(* Logix 5000 project; controller PLC_MCC1201_220AP1 vendor 1 type 14 code 164 rev 35.11; software revision 35.00; part 14 of 25 *)
(* tags used below, declared in another part *)
   AFI : ALIAS FOR B3[7].15;
   B175 : DINT[1];
   B176 : DINT[1];
   B180 : DINT[10];
   B3 : DINT[102];
   B52 : DINT[100];
   C183 : COUNTER[3];
   C1_ACTIVE_LAMP : ALIAS FOR N54[260].0;
   C2_ACTIVE_LAMP : ALIAS FOR N54[261].0;
   C3_ACTIVE_LAMP : ALIAS FOR N54[262].0;
   C5 : COUNTER[100];
   C5_ACTIVE_LAMP : ALIAS FOR N54[264].0;
   CR1_DOWN_PROX : ALIAS FOR I[64].11;
   I : INT[128];
   LEHR_2IN_PULSE : ALIAS FOR B73[0].1;
   LEHR_SPEED : ALIAS FOR N60[1];
   LEHRSPD_CURRENT : ALIAS FOR N98[5];
   MS_ACCUM : ALIAS FOR N70[1];
   MS_LEHR : ALIAS FOR N60[11];
   MSEC_TRIM : ALIAS FOR N60[12];
   N125 : DINT[414];
   N126 : DINT[103];
   N127 : DINT[997];
   N128 : DINT[997];
   N177 : DINT[5];
   N177_0 : ALIAS FOR N177[0];
   N188 : DINT[500];
   N26 : DINT[1000];
   N54 : DINT[501];
   N70 : DINT[3];
   N80 : DINT[16];
   O : INT[128];
   RELDR_ESTOP : ALIAS FOR I[80].0;
   S : INT[128];
   T182 : TIMER[11];
   T4 : TIMER[100];
   TMP_xAlwaysOFF : BOOL;
   TONY : ALIAS FOR B3[10].15;
   TRIM_2IN_PULSE : ALIAS FOR B73[0].2;
   TRIM_SPEED : ALIAS FOR N60[2];
(* MainProgram, continued *)

ROUTINE _16_PULSER   (* ladder *)
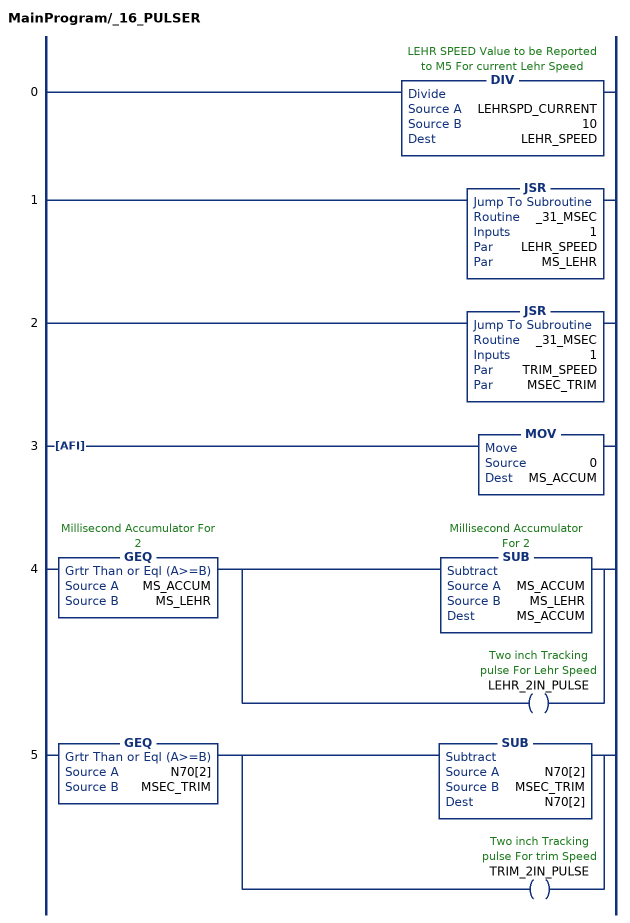
   0: DIV(LEHRSPD_CURRENT,10,LEHR_SPEED);
   1: JSR(_31_MSEC,1,LEHR_SPEED,MS_LEHR);
   2: JSR(_31_MSEC,1,TRIM_SPEED,MSEC_TRIM);
   3: AFI()MOV(0,MS_ACCUM);
   4: GEQ(MS_ACCUM,MS_LEHR)[SUB(MS_ACCUM,MS_LEHR,MS_ACCUM) ,OTE(LEHR_2IN_PULSE) ];
   5: GEQ(N70[2],MSEC_TRIM)[SUB(N70[2],MSEC_TRIM,N70[2]) ,OTE(TRIM_2IN_PULSE) ];
END_ROUTINE

ROUTINE _17_LADDER   (* ladder *)
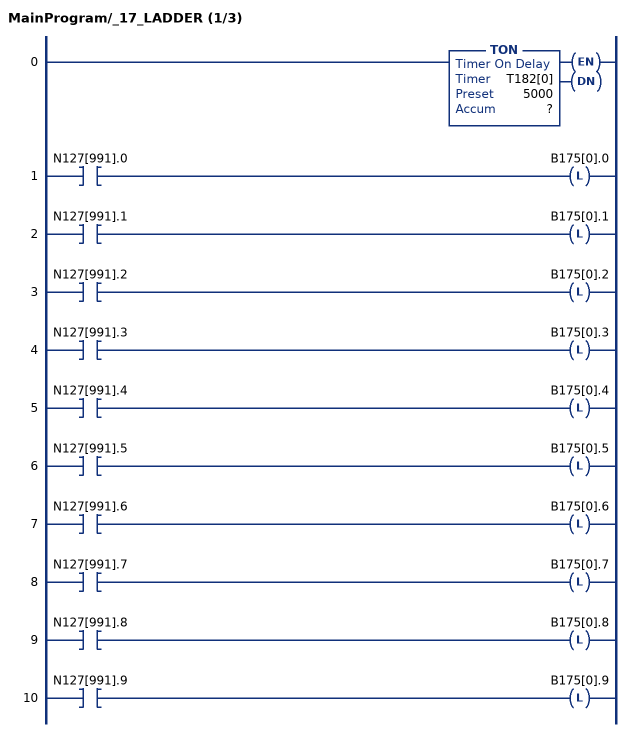
   0: TON(T182[0],?,?);
   1: XIC(N127[991].0)OTL(B175[0].0);
   2: XIC(N127[991].1)OTL(B175[0].1);
   3: XIC(N127[991].2)OTL(B175[0].2);
   4: XIC(N127[991].3)OTL(B175[0].3);
   5: XIC(N127[991].4)OTL(B175[0].4);
   6: XIC(N127[991].5)OTL(B175[0].5);
   7: XIC(N127[991].6)OTL(B175[0].6);
   8: XIC(N127[991].7)OTL(B175[0].7);
   9: XIC(N127[991].8)OTL(B175[0].8);
   10: XIC(N127[991].9)OTL(B175[0].9);
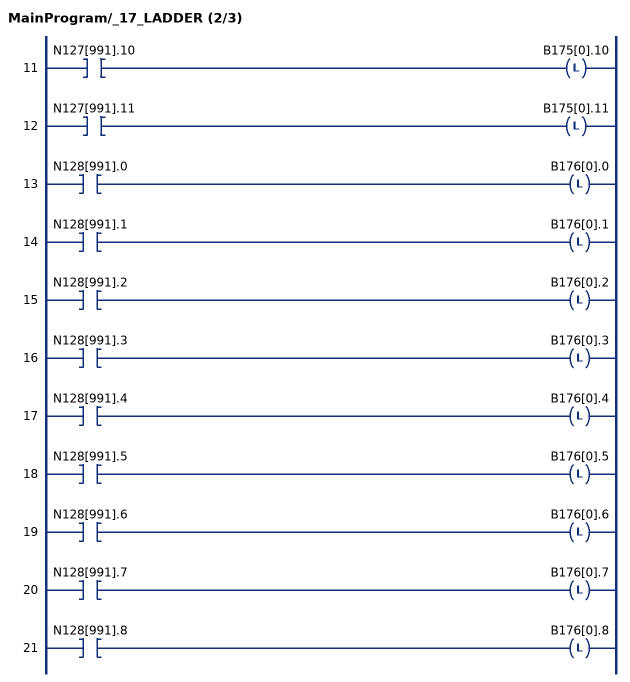
   11: XIC(N127[991].10)OTL(B175[0].10);
   12: XIC(N127[991].11)OTL(B175[0].11);
   13: XIC(N128[991].0)OTL(B176[0].0);
   14: XIC(N128[991].1)OTL(B176[0].1);
   15: XIC(N128[991].2)OTL(B176[0].2);
   16: XIC(N128[991].3)OTL(B176[0].3);
   17: XIC(N128[991].4)OTL(B176[0].4);
   18: XIC(N128[991].5)OTL(B176[0].5);
   19: XIC(N128[991].6)OTL(B176[0].6);
   20: XIC(N128[991].7)OTL(B176[0].7);
   21: XIC(N128[991].8)OTL(B176[0].8);
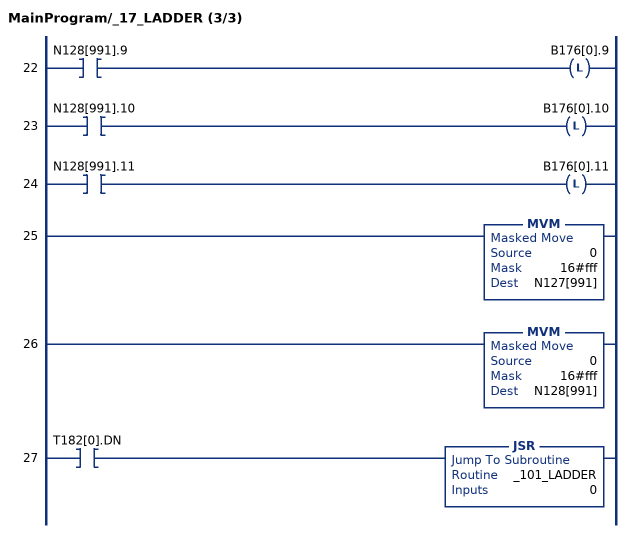
   22: XIC(N128[991].9)OTL(B176[0].9);
   23: XIC(N128[991].10)OTL(B176[0].10);
   24: XIC(N128[991].11)OTL(B176[0].11);
   25: MVM(0,16#fff,N127[991]);
   26: MVM(0,16#fff,N128[991]);
   27: XIC(T182[0].DN)JSR(_101_LADDER,0);
END_ROUTINE

ROUTINE _19_PII   (* ladder *)
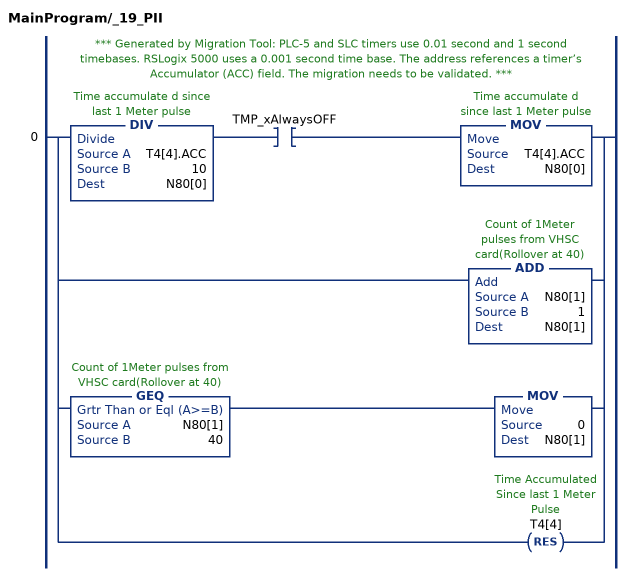
   // *** Generated by Migration Tool: PLC-5 and SLC timers use 0.01 second and 1 second timebases. RSLogix 5000 uses a 0.001 second time base. The address references a timer’s Accumulator (ACC) field. The migration needs to be validated. ***
   0: [DIV(T4[4].ACC,10,N80[0]) XIC(TMP_xAlwaysOFF) MOV(T4[4].ACC,N80[0]) ,ADD(N80[1],1,N80[1]) ,GEQ(N80[1],40) MOV(0,N80[1]) ,RES(T4[4]) ];
END_ROUTINE

ROUTINE _22_LADDER   (* ladder *)
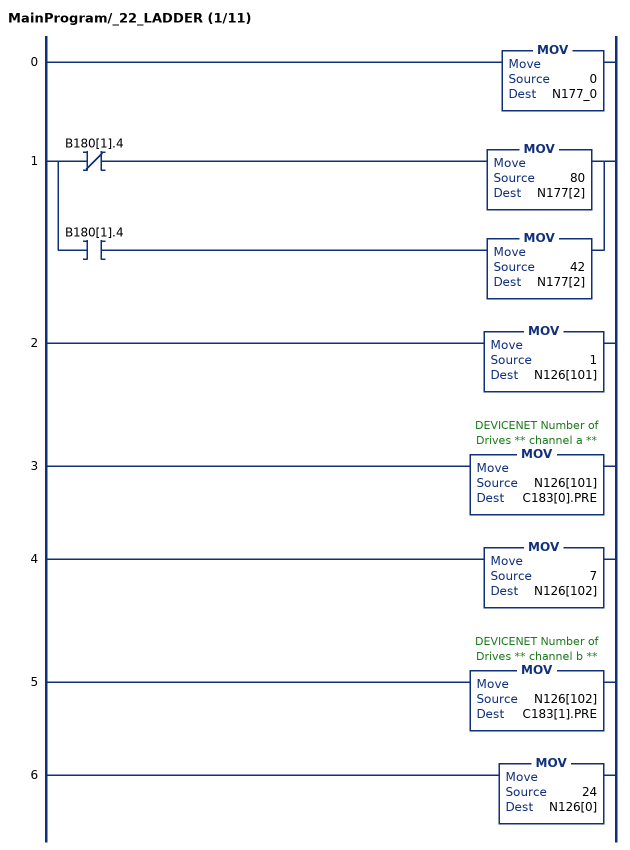
   0: MOV(0,N177_0);
   1: [XIO(B180[1].4) MOV(80,N177[2]) ,XIC(B180[1].4) MOV(42,N177[2]) ];
   2: MOV(1,N126[101]);
   3: MOV(N126[101],C183[0].PRE);
   4: MOV(7,N126[102]);
   5: MOV(N126[102],C183[1].PRE);
   6: MOV(24,N126[0]);
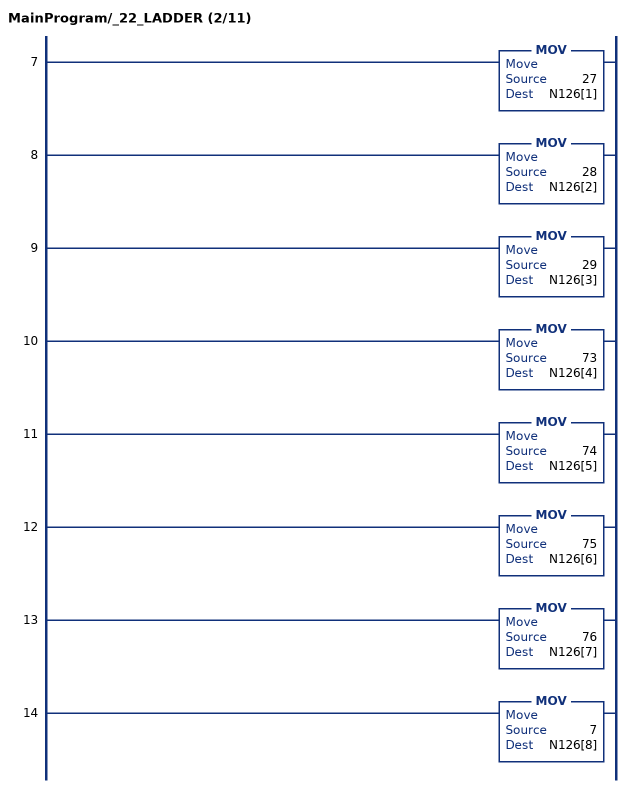
   7: MOV(27,N126[1]);
   8: MOV(28,N126[2]);
   9: MOV(29,N126[3]);
   10: MOV(73,N126[4]);
   11: MOV(74,N126[5]);
   12: MOV(75,N126[6]);
   13: MOV(76,N126[7]);
   14: MOV(7,N126[8]);
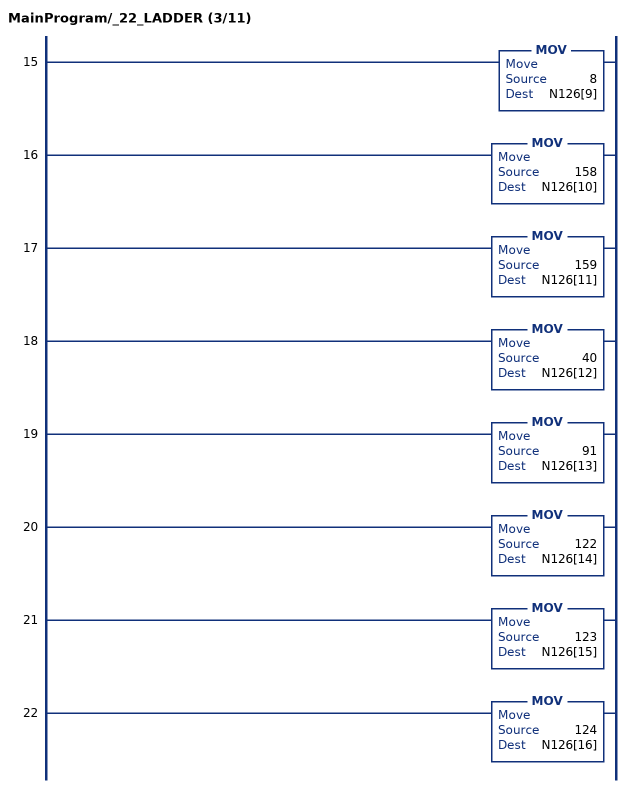
   15: MOV(8,N126[9]);
   16: MOV(158,N126[10]);
   17: MOV(159,N126[11]);
   18: MOV(40,N126[12]);
   19: MOV(91,N126[13]);
   20: MOV(122,N126[14]);
   21: MOV(123,N126[15]);
   22: MOV(124,N126[16]);
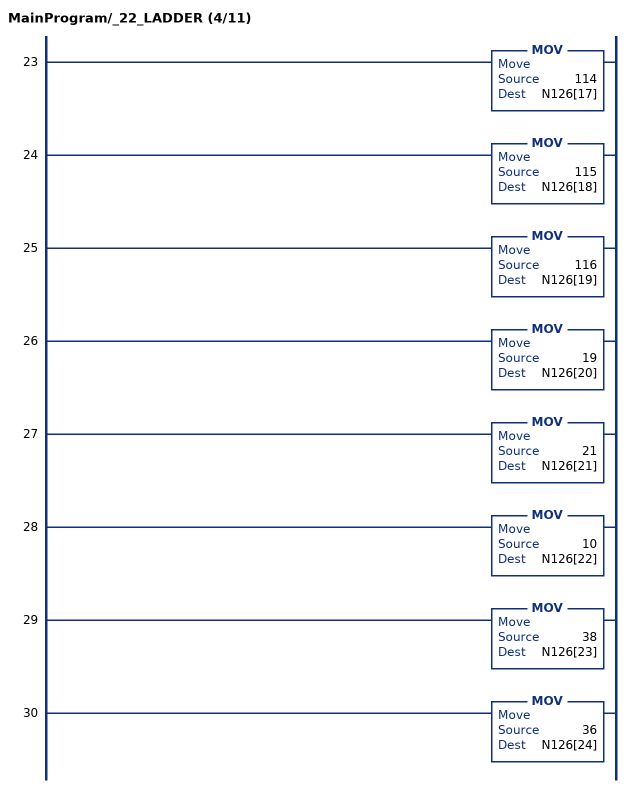
   23: MOV(114,N126[17]);
   24: MOV(115,N126[18]);
   25: MOV(116,N126[19]);
   26: MOV(19,N126[20]);
   27: MOV(21,N126[21]);
   28: MOV(10,N126[22]);
   29: MOV(38,N126[23]);
   30: MOV(36,N126[24]);
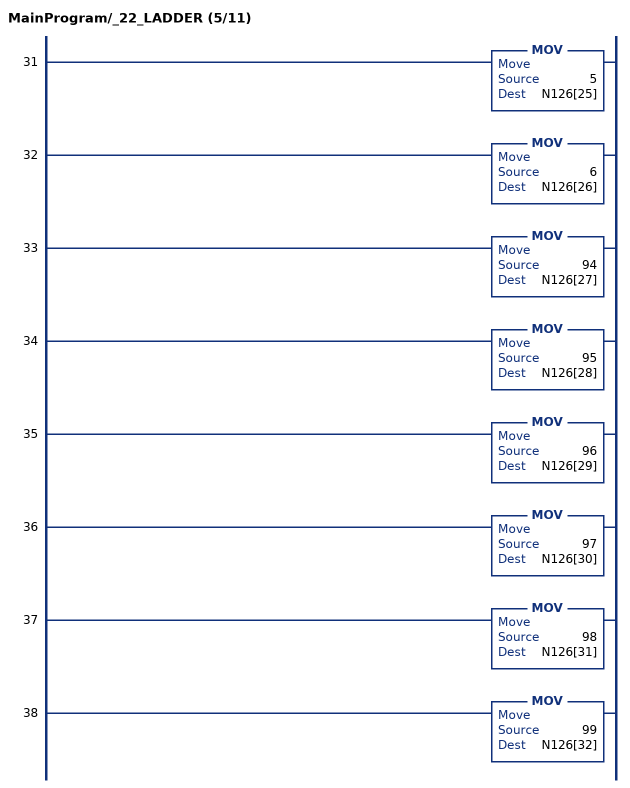
   31: MOV(5,N126[25]);
   32: MOV(6,N126[26]);
   33: MOV(94,N126[27]);
   34: MOV(95,N126[28]);
   35: MOV(96,N126[29]);
   36: MOV(97,N126[30]);
   37: MOV(98,N126[31]);
   38: MOV(99,N126[32]);
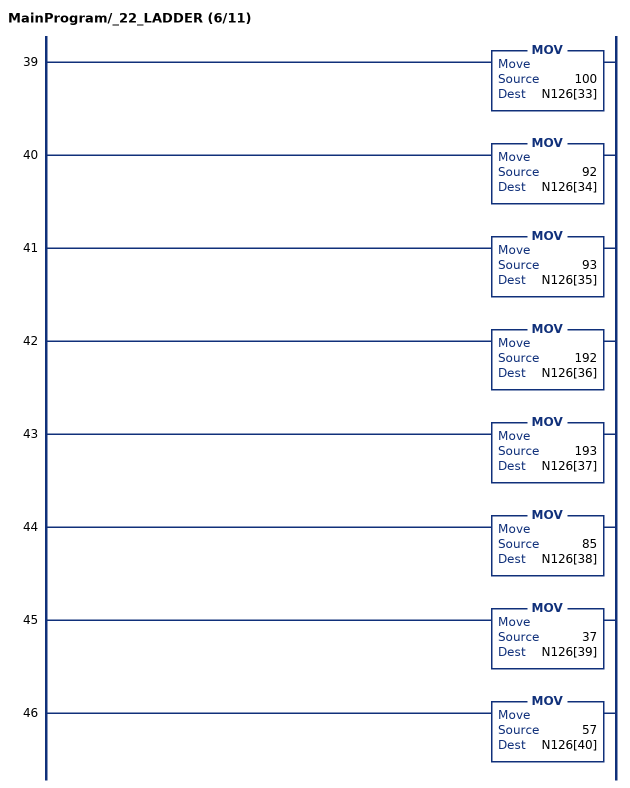
   39: MOV(100,N126[33]);
   40: MOV(92,N126[34]);
   41: MOV(93,N126[35]);
   42: MOV(192,N126[36]);
   43: MOV(193,N126[37]);
   44: MOV(85,N126[38]);
   45: MOV(37,N126[39]);
   46: MOV(57,N126[40]);
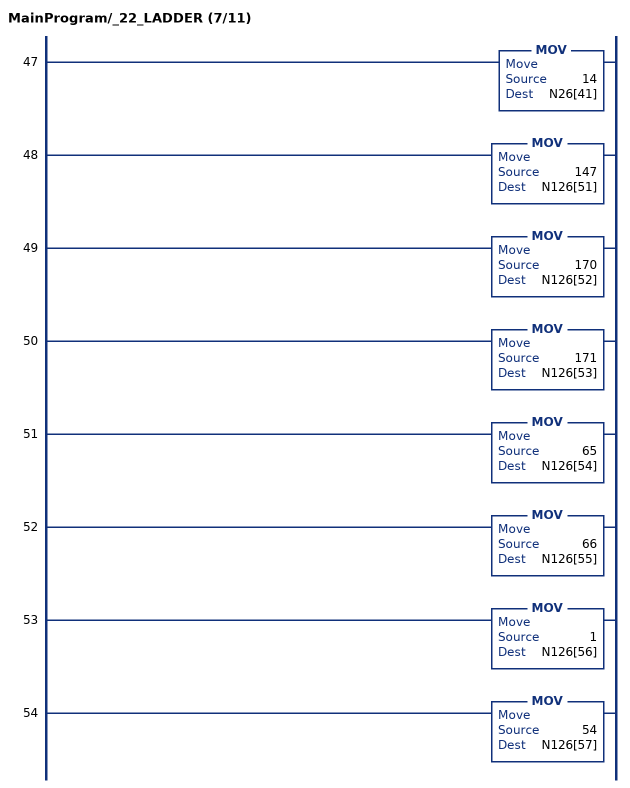
   47: MOV(14,N26[41]);
   48: MOV(147,N126[51]);
   49: MOV(170,N126[52]);
   50: MOV(171,N126[53]);
   51: MOV(65,N126[54]);
   52: MOV(66,N126[55]);
   53: MOV(1,N126[56]);
   54: MOV(54,N126[57]);
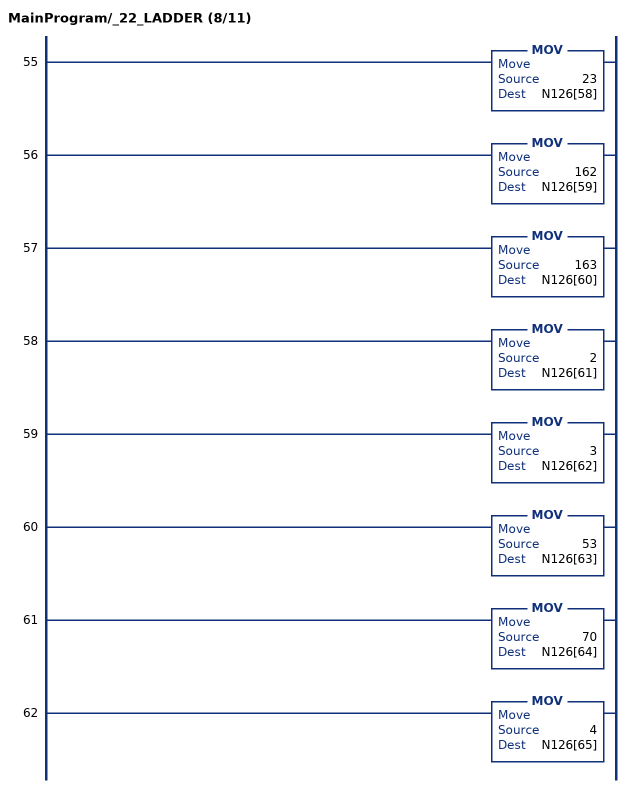
   55: MOV(23,N126[58]);
   56: MOV(162,N126[59]);
   57: MOV(163,N126[60]);
   58: MOV(2,N126[61]);
   59: MOV(3,N126[62]);
   60: MOV(53,N126[63]);
   61: MOV(70,N126[64]);
   62: MOV(4,N126[65]);
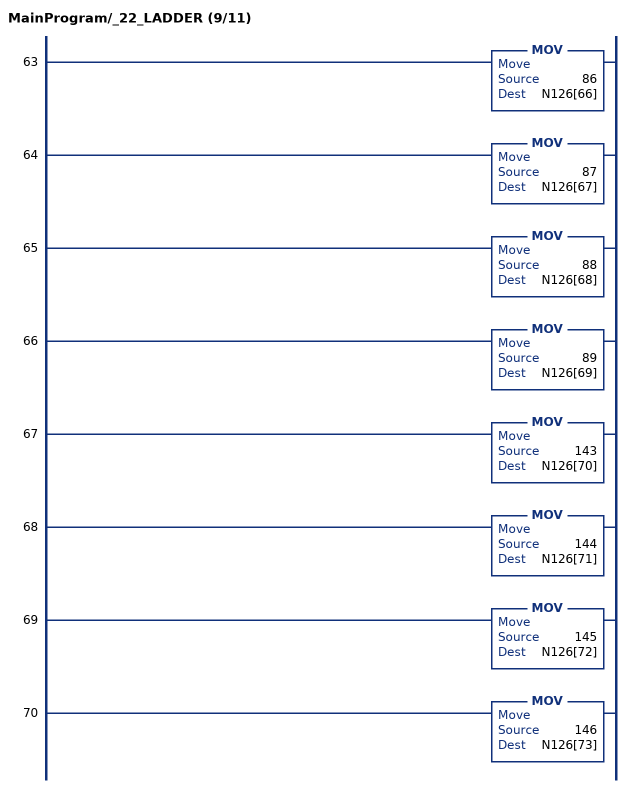
   63: MOV(86,N126[66]);
   64: MOV(87,N126[67]);
   65: MOV(88,N126[68]);
   66: MOV(89,N126[69]);
   67: MOV(143,N126[70]);
   68: MOV(144,N126[71]);
   69: MOV(145,N126[72]);
   70: MOV(146,N126[73]);
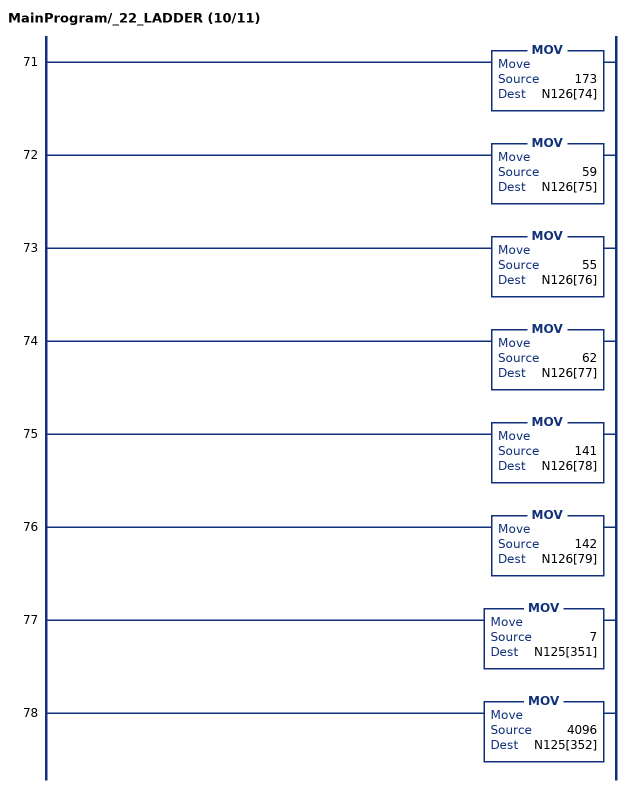
   71: MOV(173,N126[74]);
   72: MOV(59,N126[75]);
   73: MOV(55,N126[76]);
   74: MOV(62,N126[77]);
   75: MOV(141,N126[78]);
   76: MOV(142,N126[79]);
   77: MOV(7,N125[351]);
   78: MOV(4096,N125[352]);
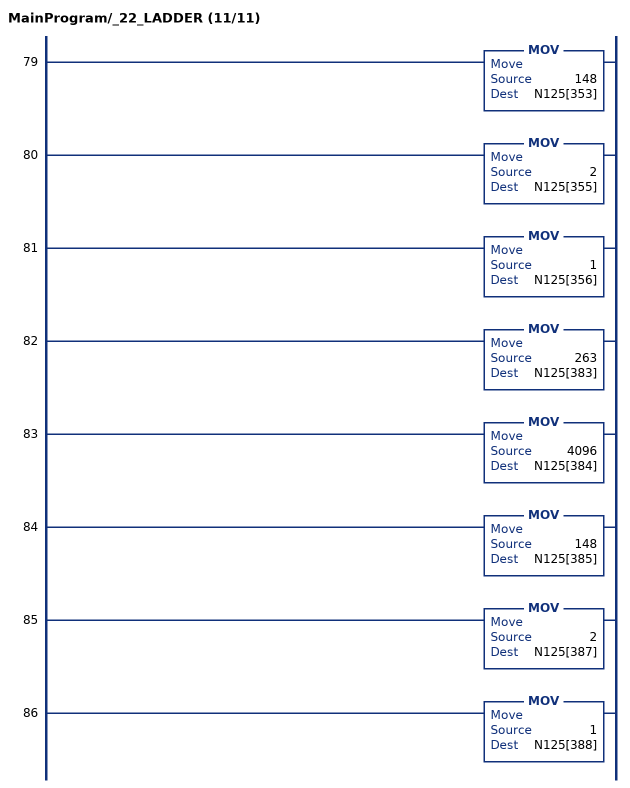
   79: MOV(148,N125[353]);
   80: MOV(2,N125[355]);
   81: MOV(1,N125[356]);
   82: MOV(263,N125[383]);
   83: MOV(4096,N125[384]);
   84: MOV(148,N125[385]);
   85: MOV(2,N125[387]);
   86: MOV(1,N125[388]);
END_ROUTINE

ROUTINE _24_ADAPTER   (* ladder *)
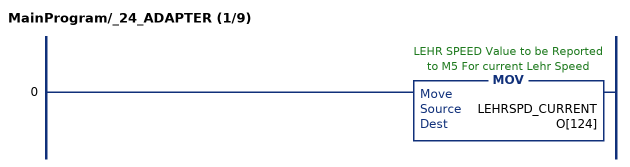
   0: MOV(LEHRSPD_CURRENT,O[124]);
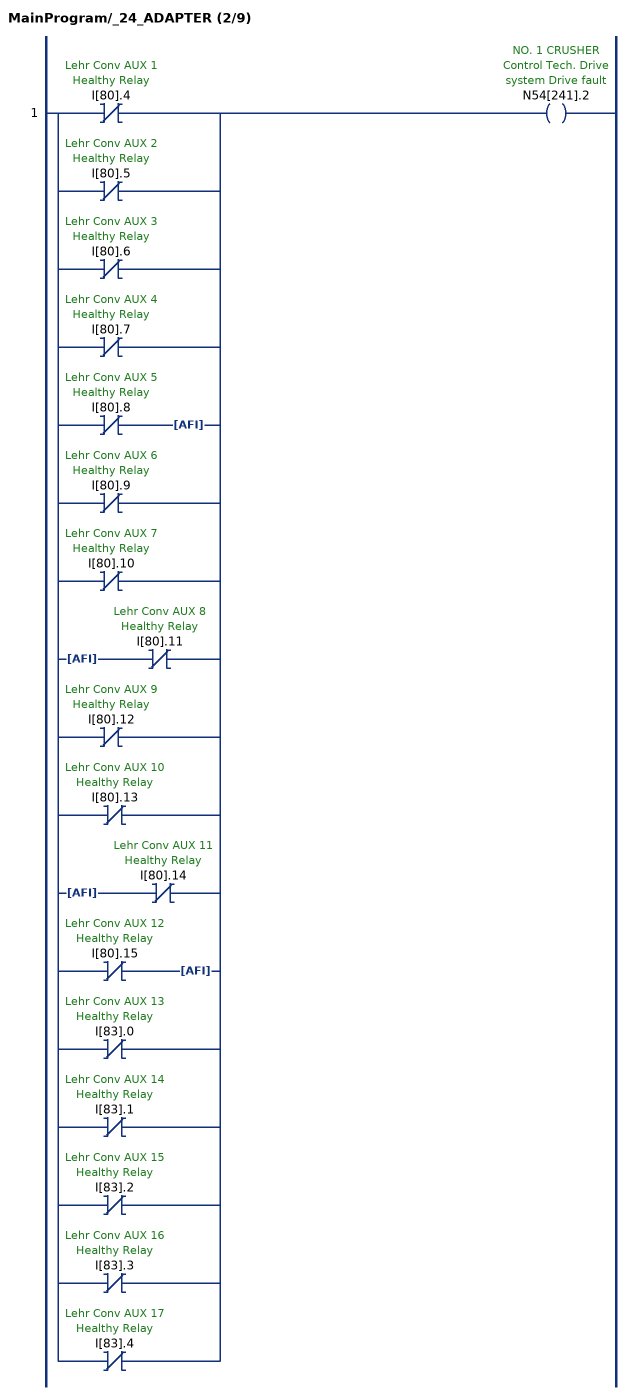
   1: [XIO(I[80].4) ,XIO(I[80].5) ,XIO(I[80].6) ,XIO(I[80].7) ,XIO(I[80].8) AFI() ,XIO(I[80].9) ,XIO(I[80].10) ,AFI() XIO(I[80].11) ,XIO(I[80].12) ,XIO(I[80].13) ,AFI() XIO(I[80].14) ,XIO(I[80].15) AFI() ,XIO(I[83].0) ,XIO(I[83].1) ,XIO(I[83].2) ,XIO(I[83].3) ,XIO(I[83].4) ]OTE(N54[241].2);
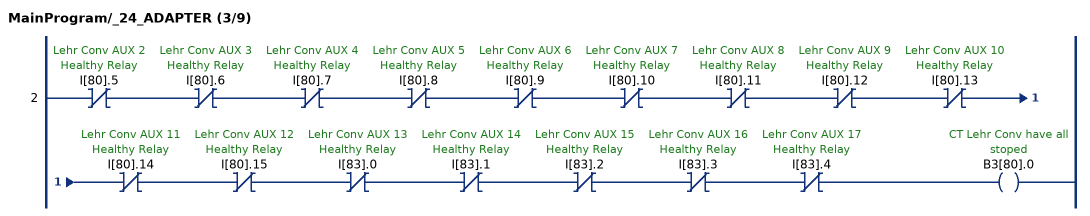
   2: XIO(I[80].5)XIO(I[80].6)XIO(I[80].7)XIO(I[80].8)XIO(I[80].9)XIO(I[80].10)XIO(I[80].11)XIO(I[80].12)XIO(I[80].13)XIO(I[80].14)XIO(I[80].15)XIO(I[83].0)XIO(I[83].1)XIO(I[83].2)XIO(I[83].3)XIO(I[83].4)OTE(B3[80].0);
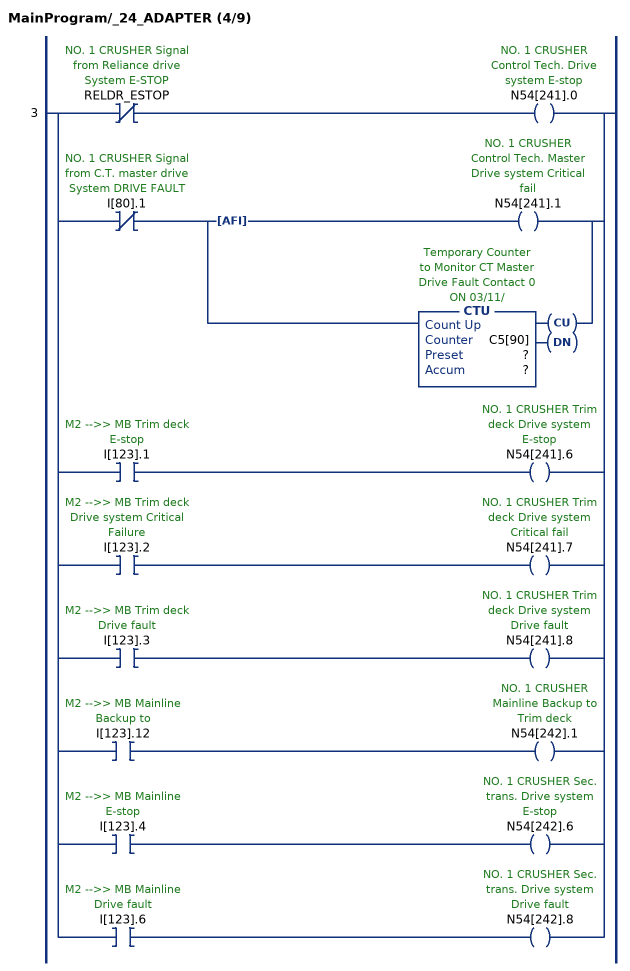
   3: [XIO(RELDR_ESTOP) OTE(N54[241].0) ,XIO(I[80].1) [AFI() OTE(N54[241].1) ,CTU(C5[90],?,?) ] ,XIC(I[123].1) OTE(N54[241].6) ,XIC(I[123].2) OTE(N54[241].7) ,XIC(I[123].3) OTE(N54[241].8) ,XIC(I[123].12) OTE(N54[242].1) ,XIC(I[123].4) OTE(N54[242].6) ,XIC(I[123].6) OTE(N54[242].8) ];
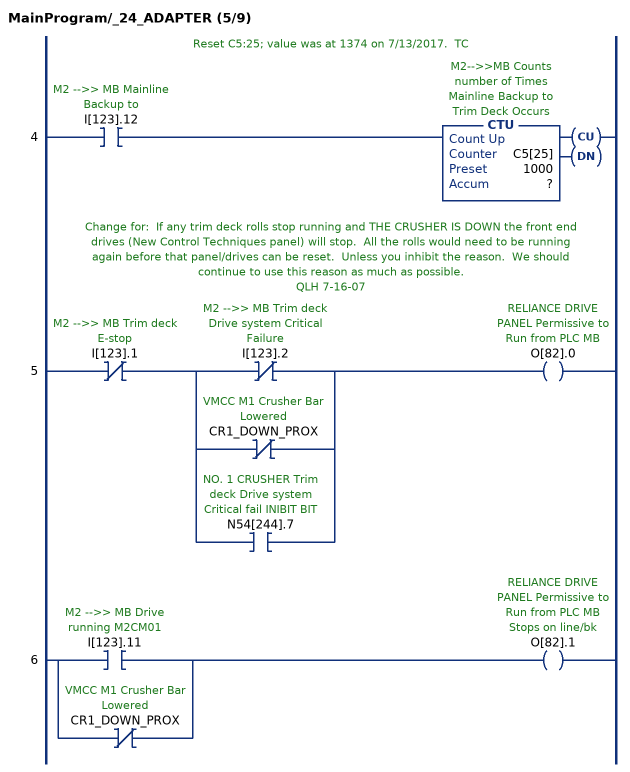
   // Reset C5:25; value was at 1374 on 7/13/2017.  TC
   4: XIC(I[123].12)CTU(C5[25],?,?);
   // Change for:  If any trim deck rolls stop running and THE CRUSHER IS DOWN the front end drives (New Control Techniques panel) will stop.  All the rolls would need to be running again before that panel/drives can be reset.  Unless you inhibit the reason.  We should continue to use this reason as much as possible.
   // QLH 7-16-07
   5: XIO(I[123].1)[XIO(I[123].2) ,XIO(CR1_DOWN_PROX) ,XIC(N54[244].7) ]OTE(O[82].0);
   6: [XIC(I[123].11) ,XIO(CR1_DOWN_PROX) ]OTE(O[82].1);
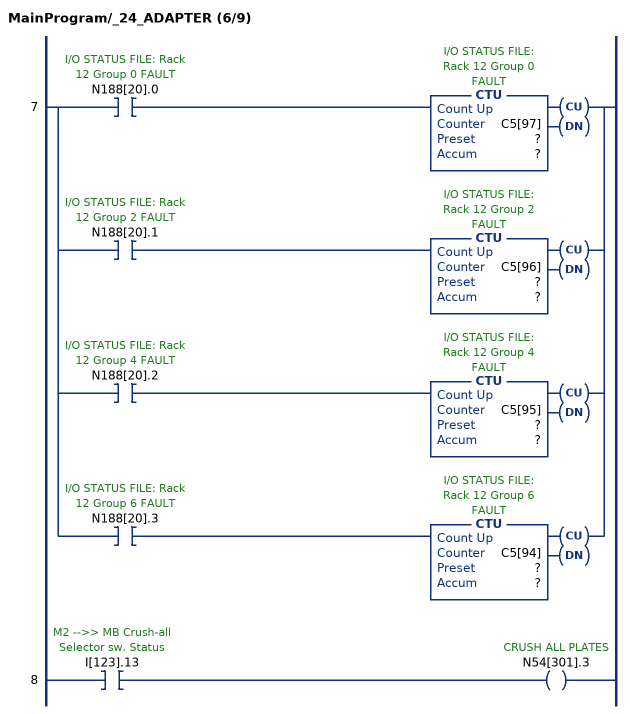
   7: [XIC(N188[20].0) CTU(C5[97],?,?) ,XIC(N188[20].1) CTU(C5[96],?,?) ,XIC(N188[20].2) CTU(C5[95],?,?) ,XIC(N188[20].3) CTU(C5[94],?,?) ];
   8: XIC(I[123].13)OTE(N54[301].3);
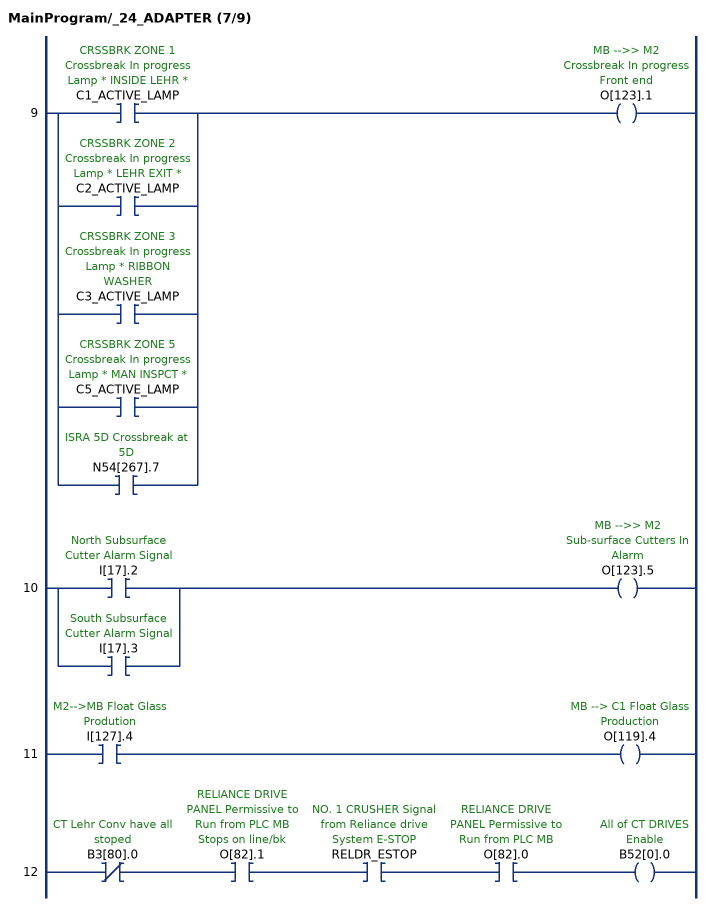
   9: [XIC(C1_ACTIVE_LAMP) ,XIC(C2_ACTIVE_LAMP) ,XIC(C3_ACTIVE_LAMP) ,XIC(C5_ACTIVE_LAMP) ,XIC(N54[267].7) ]OTE(O[123].1);
   10: [XIC(I[17].2) ,XIC(I[17].3) ]OTE(O[123].5);
   11: XIC(I[127].4)OTE(O[119].4);
   12: XIO(B3[80].0)XIC(O[82].1)XIC(RELDR_ESTOP)XIC(O[82].0)OTE(B52[0].0);
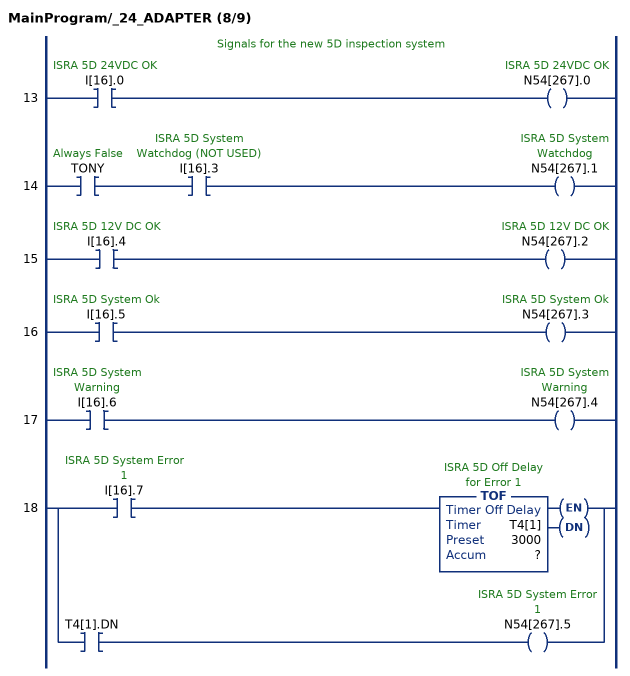
   // Signals for the new 5D inspection system
   13: XIC(I[16].0)OTE(N54[267].0);
   14: XIC(TONY)XIC(I[16].3)OTE(N54[267].1);
   15: XIC(I[16].4)OTE(N54[267].2);
   16: XIC(I[16].5)OTE(N54[267].3);
   17: XIC(I[16].6)OTE(N54[267].4);
   18: [XIC(I[16].7) TOF(T4[1],?,?) ,XIC(T4[1].DN) OTE(N54[267].5) ];
